screen "1000 - System" 1280x800, template "Top_Header"
   AlarmView "Alarm view_1" at 29,490 size 1237x294
   TextField "HmiScreenItemData" at 34,166 size 171x28; Text 'HMI device type:'
   TextField "HmiScreenItemData_5" at 240,166 size 299x28; Text 'TP1500 Comfort 15.0.1.0'
   TextField "HmiScreenItemData_7" at 34,199 size 171x28; Text 'Template Version:'
   TextField "HmiScreenItemData_8" at 34,263 size 171x28; Text 'Connection:'
   TextField "HmiScreenItemData_9" at 240,261 size 299x28; Text 'Simatic PLC Connection'
   TextField "HmiScreenItemData_10" at 34,293 size 171x28; Text 'PLC:'
   TextField "HmiScreenItemData_11" at 240,291 size 299x28; Text 'S7-1518F'
   TextField "HmiScreenItemData_1" at 240,199 size 299x28; Text 'FORD_Ver_1.1'
   TextField "HmiScreenItemData_12" at 34,231 size 171x28; Text 'Configuration Software:'
   TextField "HmiScreenItemData_13" at 240,229 size 299x28; Text 'WinCC TIA Portal V15 SP1'
   Button "HmiScreenItemData_4" at 29,119 size 283x41; TextOn 'System Information'; TextOff 'System Information'; PictureOn "Navigates to System information for TP1500 Comfort 14.0.1.0"; PictureOff "Navigates to System information for TP1500 Comfort 14.0.1.0"
   TextField "HmiScreenItemData_14" at 34,326 size 171x28; Text 'PLC Date / Time :'
   DateTimeField "Date/time field_2" at 238,356 size 253x36
   TextField "HmiScreenItemData_15" at 34,360 size 171x28; Text 'HMI Date / Time :'
   Button "HmiScreenItemData_2" at 622,114 size 262x48; TextOn 'System Settings'; TextOff 'System Settings'; PictureOn "Navigates to System settings for TP1500 Comfort 14.0.1.0"; PictureOff "Navigates to System settings for TP1500 Comfort 14.0.1.0"
   Button "HmiScreenItemData_6" at 29,442 size 318x44; TextOn 'System Messages'; TextOff 'System Messages'; PictureOn "Navigates to System screens for TP1500 Comfort 14.0.1.0"; PictureOff "Navigates to System screens for TP1500 Comfort 14.0.1.0"
      on Release: ActivateScreen("1000 - System", 0)
   TextField "Text field_1" at 241,328 size 48x31; Text 'Text'
   Button "Toggle language_1" at 1082,171 size 101x121; TextOn 'Toggle langu...'; TextOff 'User Admin.'
      on Release: ActivateScreen("1001 - User Adminstration", 0)
   Button "Toggle language_2" at 622,171 size 101x121; TextOn 'Toggle langu...'; TextOff 'Online'
      on Release: function_bb44b551(0)
   Button "Toggle language_3" at 736,171 size 101x121; TextOn 'Toggle langu...'; TextOff 'Offline'
      on Release: function_bb44b551(1)
   Button "Toggle language_4" at 851,171 size 101x121; TextOn 'Toggle langu...'; TextOff 'Transfer'
      on Release: function_bb44b551(2)
   Button "Toggle language_5" at 966,171 size 101x121; TextOn 'Toggle langu...'; TextOff 'Toggle Language'
      on Release: function_fb9197e8(-1)
   Button "Toggle language_6" at 622,301 size 101x121; TextOn 'Toggle langu...'; TextOff 'Calibrate Screen'
      on Release: function_bc3e350c()
   Button "Toggle language_7" at 736,301 size 101x121; TextOn 'Toggle langu...'; TextOff 'Clean Screen'
      on Release: function_be740847(30)
   Button "Toggle language_8" at 851,301 size 101x121; TextOn 'Toggle langu...'; TextOff 'Control Panel'
      on Release: function_f34a74f3()
   Button "Toggle language_9" at 965,301 size 101x121; TextOn 'Toggle langu...'; TextOff 'Stop Runtime'
      on Release: StopRuntime(0)
   Button "Toggle language_10" at 472,301 size 101x121; TextOn 'Toggle langu...'; TextOff 'Internal Software Versions'
      on Release: function_febcb963(-1)
   Button "Button_1" at 1082,301 size 102x120; TextOff 'On Screen Keyboard'
      on Release: function_d6caf649(0)
      Appearance <- "Always_OFF_HMI"

screen "1001 - User Adminstration" 1280x800, template "Top_Header"
   UserView "User view_1" at 26,185 size 1235x486
   Button "HmiScreenItemData_3" at 48,119 size 197x58; TextOn 'User Administration'; TextOff 'User Administration'; PictureOn "Navigates to User administration for TP1500 Comfort 14.0.1.0"; PictureOff "Navigates to User administration for TP1500 Comfort 14.0.1.0"

Template "TESTCENTER_SDC" 1280x800
   Button "Template_Vorlage_Schaltfläche" at 260,714 size 128x84; TextOff 'START'
      on Click: ActivateScreen("010_START", 0)
   Button "Template_Vorlage_Schaltfläche_0" at 387,714 size 128x84; TextOff 'OVERVIEW'
      on Click: ActivateScreen("700_System_Line_Overview", 0)
   Button "Template_Vorlage_Schaltfläche_1" at 514,714 size 128x84; TextOff 'TS PARAMETER'
      on Click: ActivateScreen("708_ZONE_STATUS", 0); "SDC_TS_PARAMETER"()
   Button "Template_Vorlage_Schaltfläche_2" at 641,714 size 128x84; TextOff 'EMS STATUS'
      on Click: ActivateScreen("711_CARRIER_STATUS", 0)
   Button "Template_Vorlage_Schaltfläche_3" at 768,714 size 128x84; TextOff 'Text'
   Button "Template_Vorlage_Schaltfläche_4" at 895,714 size 128x84; TextOff 'MESSAGES'
      on Click: ActivateScreen("019_MESSAGEs", 0)
   Button "Template_Vorlage_Schaltfläche_5" at 1022,714 size 128x84; TextOff 'FEHLER QUIT FAULT RESET'
      on Release: ResetBit("DB_SDC_GLOBAL_M.SDC_ER_Reset(1)")
      on Press: SetBit("DB_SDC_GLOBAL_M.SDC_ER_Reset(1)")
   Button "Template_Vorlage_Schaltfläche_6" at 1149,714 size 128x84; TextOff 'zurück / BACK'
      on Click: function_efd93a16()
   SymbolicIOField "Template_Vorlage_Symbolisches EA-Feld" at 1,3 size 671x25; TextOn '1'; TextOff '0'; TextList "SDC_ScreensName"
      ProcessValue <- "SDC\_intern_Bildnummer"
   UserView "Template_Vorlage_Vorlage_Benutzeranzeige_1" at 935,3 size 175x24
   DateTimeField "Template_Vorlage_DateTimeField_1" at 868,3 size 65x22
   DateTimeField "Template_Vorlage_DateTimeField_0" at 784,4 size 87x20
   GraphicView "Template_Vorlage_TemplateGraphicViewLogo_1" at 1112,3 size 167x25; Picture "Siemens"
   GraphicIOField "Template_Vorlage_Grafisches EA-Feld_1" at 2,4 size 20x20; PictureList "Grafikliste_G_Y"
      ProcessValue <- "Clock_1Hz"
   IOField "Vorlage_EA-Feld_2" at 754,4 size 44x19; FormatPattern 9999
      ProcessValue <- "_intern_Pult_Nr"
   TextField "Vorlage_Textfeld_1" at 677,3 size 89x23; Text 'PultNr. SDC'
   Button "Template_Vorlage_Schaltfläche_7" at 2,714 size 258x84; TextOff 'Text'
   AlarmView "Template_Vorlage_AlarmsLine_1" at 0,676 size 1280x36; ColumnTextDevice 'PLC / Steuerung / ПЛК'; ColumnTextNumber 'Nr. / No. / 编号 / № / N.º.'; ColumnTextAckGroup 'Gruppe quittieren / QGR / Acknowledge group / 确认组 / Квитировать группу / Acusar grupo'; ColumnTextAlarmState 'Status / Zustand / 状态 / Статус / Estado'; ColumnTextTime 'Zeit / Uhrzeit / Time / 时间 / Время / Hora'; ColumnTextDate 'Datum / Date / 日期 / Дата / Fecha'; ColumnTextAlarmText 'Text / 文本 / Текст / Texto'

Template "SDC" 1280x800
   SymbolicIOField "Template_Vorlage_Symbolisches EA-Feld" at 261,2 size 708x31; TextOn '1'; TextOff '0'; TextList "SDC_ScreensName"
      ProcessValue <- "SDC\_intern_Bildnummer"
   GraphicView "Template_Vorlage_TemplateGraphicViewLogo_1" at 1107,5 size 167x25; Picture "Siemens"
   GraphicIOField "Template_Vorlage_Grafisches EA-Feld_1" at 1081,8 size 20x20; PictureList "Grafikliste_G_Y"
      ProcessValue <- "Clock_1Hz"
   Button "Template_Vorlage_Schaltfläche" at 11,714 size 128x84; TextOff 'HOME / START'
      on Click: ActivateScreen("010_START", 0)
   Button "Template_Vorlage_Schaltfläche_1" at 271,714 size 128x84; TextOff 'TS PAR. TS PARAMETER'
      on Click: ActivateScreen("708_ZONE_STATUS", 0); "SDC_TS_PARAMETER"()
   Button "Template_Vorlage_Schaltfläche_2" at 401,714 size 128x84; TextOff 'EMS STATUS'
      on Click: ActivateScreen("711_CARRIER_STATUS", 0)
   Button "Template_Vorlage_Schaltfläche_4" at 888,714 size 128x84; TextOff 'ERRORS / MESSAGES / MELDUNGEN'
      on Click: ActivateScreen("019_MESSAGEs", 0)
   Button "Template_Vorlage_Schaltfläche_5" at 1018,714 size 128x84; TextOff 'QUIT FAULT RESET'
      on Release: ResetBit("DB_SDC_GLOBAL_M.SDC_ER_Reset")
      on Press: SetBit("DB_SDC_GLOBAL_M.SDC_ER_Reset")
   Button "Template_Vorlage_Schaltfläche_6" at 1148,714 size 128x84; TextOff 'BACK / ZURÜCK'
      on Click: function_efd93a16()
   Button "Template_Vorlage_Schaltfläche_3" at 141,714 size 128x84; TextOff 'GLOB. PAR. START GLOBAL PARAMETER'
      on Click: ActivateScreen("707_GLOBAL_PARAMETER", 0)
   TextField "Vorlage_Textfeld_1" at 909,6 size 127x25; Text 'DeskNo. SDC'
   IOField "Vorlage_EA-Feld_1" at 1039,4 size 41x29; FormatPattern 999
      ProcessValue <- "_intern_Pult_Nr"
   TextField "Template_Vorlage_OBJECT_3" at 1,1 size 70x32; Text 'TIME: / Zeit:'
      Appearance <- "TP_Online"
   DateTimeField "Template_Vorlage_OBJECT_5" at 56,1 size 114x32
      Appearance <- "TP_Online"
   DateTimeField "Vorlage_Datum/Uhrzeit-Feld_1" at 169,4 size 123x26

Template "Top_Header" 1280x800
   Button "Template_Button_3" at 1074,2 size 203x55; TextOn 'FAULT RESET FAULT RESET'; TextOff 'FAULT RESET FAULT RESET'
      on Release: ResetBit("DB_SDC_GLOBAL_M.SDC_ER_Reset")
      on Press: SetBit("DB_SDC_GLOBAL_M.SDC_ER_Reset")
   AlarmView "Template_Alarm view_2" at 128,2 size 948x112
   Button "Template_Button_4" at 1196,56 size 81x59; TextOff 'Text'
      Appearance <- "AlwaysTRUE"
   Button "Button_7" at 0,57 size 128x58; TextOff 'SELECT SCREEN'
      on Release: ActivateScreen("010_START", 0)
   Button "Button_6" at 0,0 size 128x58; TextOff 'PREVIOUS SCREEN'
      on Click: function_efd93a16()
   DateTimeField "Template_Date/time field_2" at 1075,56 size 123x28
   DateTimeField "Template_Date/time field_3" at 1075,83 size 122x32

PopupScreen "Pop-up_OverviewModules" 1280x800
   Button "Schaltfläche_64" at 1110,723 size 119x49; TextOn 'schließen / close'; TextOff 'schließen / close'
      on Click: function_efd93a16("Pop-up_OverviewModules", 0, 0, 0, -1, 2); ResetBit("UserDiag_HmiData_ioSlotDiagnosticsLoaded")
   IOField "I/O field_2" at 241,713 size 579x49; FormatPattern ??????????????????????????????????????????????????
      ProcessValue <- "UserDiag_HmiData_actDeviceName"
   IOField "I/O field_1" at 241,647 size 60x49; FormatPattern 999
      ProcessValue <- "actIOSystemNumber"
   IOField "I/O field_3" at 383,647 size 60x49; FormatPattern 999
      ProcessValue <- "UserDiag_HmiData_actDeviceNumber"
   TextField "Text field_1" at 137,658 size 107x26; Text 'IO System'
   TextField "Text field_2" at 314,658 size 72x26; Text 'Device'
      Visibility <- "actIOSystemNumber"
   TextField "Text field_3" at 181,724 size 62x26; Text 'Name'
   ScreenModuleView "typeSlot_1" at 67,22 size 49x152; Guid_{11997190-58737} '01'; ScreenModuleType ""
      Guid_{11997190-58740} <- "[1]"
      Guid_{11997190-58743} <- "[1]"
   ScreenModuleView "typeSlot_2" at 20,22 size 49x152; ScreenModuleType ""
      Guid_{11997190-58740} <- "[0]"
      Guid_{11997190-58743} <- "[0]"
   ScreenModuleView "typeSlot_3" at 115,22 size 49x152; Guid_{11997190-58737} '02'; ScreenModuleType ""
      Guid_{11997190-58740} <- "[2]"
      Guid_{11997190-58743} <- "[2]"
   ScreenModuleView "typeSlot_4" at 162,22 size 49x152; Guid_{11997190-58737} '03'; ScreenModuleType ""
      Guid_{11997190-58740} <- "[3]"
      Guid_{11997190-58743} <- "[3]"
   ScreenModuleView "typeSlot_5" at 210,22 size 49x152; Guid_{11997190-58737} '04'; ScreenModuleType ""
      Guid_{11997190-58740} <- "[4]"
      Guid_{11997190-58743} <- "[4]"
   ScreenModuleView "typeSlot_6" at 257,22 size 49x152; Guid_{11997190-58737} '05'; ScreenModuleType ""
      Guid_{11997190-58740} <- "[5]"
      Guid_{11997190-58743} <- "[5]"
   ScreenModuleView "typeSlot_7" at 305,22 size 49x152; Guid_{11997190-58737} '06'; ScreenModuleType ""
      Guid_{11997190-58740} <- "[6]"
      Guid_{11997190-58743} <- "[6]"
   ScreenModuleView "typeSlot_8" at 352,22 size 49x152; Guid_{11997190-58737} '07'; ScreenModuleType ""
      Guid_{11997190-58740} <- "[7]"
      Guid_{11997190-58743} <- "[7]"
   ScreenModuleView "typeSlot_9" at 400,22 size 49x152; Guid_{11997190-58737} '08'; ScreenModuleType ""
      Guid_{11997190-58740} <- "[8]"
      Guid_{11997190-58743} <- "[8]"
   ScreenModuleView "typeSlot_10" at 447,22 size 49x152; Guid_{11997190-58737} '09'; ScreenModuleType ""
      Guid_{11997190-58740} <- "[9]"
      Guid_{11997190-58743} <- "[9]"
   ScreenModuleView "typeSlot_11" at 495,22 size 49x152; Guid_{11997190-58737} '10'; ScreenModuleType ""
      Guid_{11997190-58740} <- "[10]"
      Guid_{11997190-58743} <- "[10]"
   ScreenModuleView "typeSlot_12" at 542,22 size 49x152; Guid_{11997190-58737} '11'; ScreenModuleType ""
      Guid_{11997190-58740} <- "[11]"
      Guid_{11997190-58743} <- "[11]"
   ScreenModuleView "typeSlot_13" at 590,22 size 49x152; Guid_{11997190-58737} '12'; ScreenModuleType ""
      Guid_{11997190-58740} <- "[12]"
      Guid_{11997190-58743} <- "[12]"
   ScreenModuleView "typeSlot_14" at 637,22 size 49x152; Guid_{11997190-58737} '13'; ScreenModuleType ""
      Guid_{11997190-58740} <- "[13]"
      Guid_{11997190-58743} <- "[13]"
   ScreenModuleView "typeSlot_15" at 685,22 size 49x152; Guid_{11997190-58737} '14'; ScreenModuleType ""
      Guid_{11997190-58740} <- "[14]"
      Guid_{11997190-58743} <- "[14]"
   ScreenModuleView "typeSlot_16" at 733,22 size 49x152; Guid_{11997190-58737} '15'; ScreenModuleType ""
      Guid_{11997190-58740} <- "[15]"
      Guid_{11997190-58743} <- "[15]"
   ScreenModuleView "typeSlot_17" at 780,22 size 49x152; Guid_{11997190-58737} '16'; ScreenModuleType ""
      Guid_{11997190-58740} <- "[16]"
      Guid_{11997190-58743} <- "[16]"
   ScreenModuleView "typeSlot_18" at 828,22 size 49x152; Guid_{11997190-58737} '17'; ScreenModuleType ""
      Guid_{11997190-58740} <- "[17]"
      Guid_{11997190-58743} <- "[17]"
   ScreenModuleView "typeSlot_19" at 875,22 size 49x152; Guid_{11997190-58737} '18'; ScreenModuleType ""
      Guid_{11997190-58740} <- "[18]"
      Guid_{11997190-58743} <- "[18]"
   ScreenModuleView "typeSlot_20" at 923,22 size 49x152; Guid_{11997190-58737} '19'; ScreenModuleType ""
      Guid_{11997190-58740} <- "[19]"
      Guid_{11997190-58743} <- "[19]"
   ScreenModuleView "typeSlot_21" at 971,22 size 49x152; Guid_{11997190-58737} '20'; ScreenModuleType ""
      Guid_{11997190-58740} <- "[20]"
      Guid_{11997190-58743} <- "[20]"
   ScreenModuleView "typeSlot_22" at 20,197 size 49x152; Guid_{11997190-58737} '21'; ScreenModuleType ""
      Guid_{11997190-58740} <- "[21]"
      Guid_{11997190-58743} <- "[21]"
   ScreenModuleView "typeSlot_23" at 67,197 size 49x152; Guid_{11997190-58737} '22'; ScreenModuleType ""
      Guid_{11997190-58740} <- "[22]"
      Guid_{11997190-58743} <- "[22]"
   ScreenModuleView "typeSlot_24" at 115,197 size 49x152; Guid_{11997190-58737} '23'; ScreenModuleType ""
      Guid_{11997190-58740} <- "[23]"
      Guid_{11997190-58743} <- "[23]"
   ScreenModuleView "typeSlot_25" at 162,197 size 49x152; Guid_{11997190-58737} '24'; ScreenModuleType ""
      Guid_{11997190-58740} <- "[24]"
      Guid_{11997190-58743} <- "[24]"
   ScreenModuleView "typeSlot_26" at 210,197 size 49x152; Guid_{11997190-58737} '25'; ScreenModuleType ""
      Guid_{11997190-58740} <- "[25]"
      Guid_{11997190-58743} <- "[25]"
   ScreenModuleView "typeSlot_27" at 257,197 size 49x152; Guid_{11997190-58737} '26'; ScreenModuleType ""
      Guid_{11997190-58740} <- "[26]"
      Guid_{11997190-58743} <- "[26]"
   ScreenModuleView "typeSlot_28" at 305,197 size 49x152; Guid_{11997190-58737} '27'; ScreenModuleType ""
      Guid_{11997190-58740} <- "[27]"
      Guid_{11997190-58743} <- "[27]"
   ScreenModuleView "typeSlot_29" at 352,197 size 49x152; Guid_{11997190-58737} '28'; ScreenModuleType ""
      Guid_{11997190-58740} <- "[28]"
      Guid_{11997190-58743} <- "[28]"
   ScreenModuleView "typeSlot_30" at 400,197 size 49x152; Guid_{11997190-58737} '29'; ScreenModuleType ""
      Guid_{11997190-58740} <- "[29]"
      Guid_{11997190-58743} <- "[29]"
   ScreenModuleView "typeSlot_31" at 448,197 size 49x152; Guid_{11997190-58737} '30'; ScreenModuleType ""
      Guid_{11997190-58740} <- "[30]"
      Guid_{11997190-58743} <- "[30]"
   ScreenModuleView "typeSlot_32" at 495,197 size 49x152; Guid_{11997190-58737} '31'; ScreenModuleType ""
      Guid_{11997190-58740} <- "[31]"
      Guid_{11997190-58743} <- "[31]"
   IOField "I/O field_4" at 562,647 size 60x49; FormatPattern 999
      Visibility <- "actIOSystemNumber"
      ProcessValue <- "[0]"
   TextField "Text field_4" at 452,658 size 112x26; Text 'IP Adresse / IP address'
      Visibility <- "actIOSystemNumber"
   IOField "I/O field_5" at 628,647 size 60x49; FormatPattern 999
      Visibility <- "actIOSystemNumber"
      ProcessValue <- "[1]"
   IOField "I/O field_6" at 694,647 size 60x49; FormatPattern 999
      Visibility <- "actIOSystemNumber"
      ProcessValue <- "[2]"
   IOField "I/O field_7" at 760,647 size 60x49; FormatPattern 999
      Visibility <- "actIOSystemNumber"
      ProcessValue <- "[3]"
   TextField "Text field_5" at 325,658 size 58x26; Text 'Slave'
      Visibility <- "actIOSystemNumber"

PopupScreen "Pop-up_Legend" 1280x800
   TextField "Text field_1" at 15,5 size 100x49; Text 'Legende / Legend'
   TextField "Text field_2" at 80,80 size 103x26; Text 'Status OK / State OK'
   TextField "Text field_3" at 80,146 size 165x26; Text 'Status GESTÖRT / State FAULTY'
   TextField "Text field_4" at 80,212 size 254x26; Text 'Status AUSGEFALLEN / State LOST CONNECTION'
   TextField "Text field_5" at 80,277 size 211x26; Text 'Status DEAKTIVIERT / State DEACTIVATED'
   TextField "Text field_6" at 80,343 size 339x26; Text 'Status PROBLEM / MAINTENANCE / State PROBLEM / MAINTENANCE'
   TextField "Text field_7" at 80,409 size 268x26; Text 'Status GESTÖRT GEWESEN / State WAS FAULTY'
   TextField "Text field_8" at 80,475 size 315x26; Text 'Status AUSGEFALLEN GEWESEN / State HAD LOST CONNECTION'
   TextField "Text field_9" at 80,540 size 314x26; Text 'Status DEAKTIVIERT GEWESEN / State WAS DEACTIVATED'
   TextField "Text field_10" at 80,606 size 442x26; Text 'Status PROBLEM / MAINTENANCE GEWESEN / State WAS PROBLEM / MAINTENANCE'
   Button "Schaltfläche_64" at 1110,723 size 119x49; TextOn 'schließen / close'; TextOff 'schließen / close'
      on Click: function_efd93a16("Pop-up_Legend", 0, 0, 0, -1, 2)

screen "010_START" 1280x800, template "Top_Header"
   on GenerateScreen: function_ea909784(0, U 0, '\Storage Card USB\record.csv', 2, 1, N)
   Button "Button_1" at 775,328 size 140x105; TextOn 'GLOBAL_PARAMETER GLOBAL PARAMETER'; TextOff 'GLOBAL_PARAMETER GLOBAL PARAMETER'
      on Click: ActivateScreen("707_GLOBAL_PARAMETER", 0)
   Button "Button_7" at 535,327 size 140x105; TextOn 'SECTION STATUS SECTION STATUS'; TextOff 'SECTION STATUS ZONE STATUS'
      on Click: ActivateScreen("708_ZONE_STATUS", 0)
   Button "Button_9" at 535,454 size 140x105; TextOn 'EMS STATUS EMS STATUS'; TextOff 'EMS STATUS CARRIER STATUS'
      on Click: ActivateScreen("711_CARRIER_STATUS", 0)
   Button "Button_14" at 535,198 size 140x105; TextOn 'LINE_OVERVIEW_2 LINE OVERVIEW_2'; TextOff 'LINE_OVERVIEW_2 LINE OVERVIEW'
      on Click: ActivateScreen("700_System_Line_Overview", 0)
   Button "Button_17" at 775,585 size 140x105; TextOn 'LINE_OVERVIEW_1 / MESSAGES'; TextOff 'LINE_OVERVIEW_1 FAULT MESSAGES'
      on Click: ActivateScreen("019_MESSAGEs", 0)
   Button "Button_18" at 775,454 size 140x105; TextOn 'LINE_OVERVIEW_1 PROFINET IO DIAGNOSTICS'; TextOff 'LINE_OVERVIEW_1 PROFINET IO DIAGNOSTICS'
      on Click: ActivateScreen("752_Profinet_IO_System", 0)
   Button "Button_3" at 535,585 size 140x105; TextOn 'EMS STATUS EMS STATUS'; TextOff 'EMS STATUS ALL CARRIER STATUS'
      on Click: ActivateScreen("710_ALL_CARRIER_STATUS", 0)
   Button "Button_6" at 299,198 size 140x105; TextOn 'SECTION PARAMETER SECTION PARAMETER'; TextOff 'SECTION PARAMETER SYSTEM SCREEN'
      on Click: ActivateScreen("1000 - System", 0)
   Button "Button_10" at 299,323 size 140x105; TextOn 'SECTION STATUS SECTION STATUS'; TextOff 'SECTION STATUS SYSTEM DIAGNOSTIC'
      on Release: ActivateScreen("2003 - System Diag", 0)
   Button "Button_12" at 299,450 size 140x105; TextOn 'SECTION STATUS SECTION STATUS'; TextOff 'SECTION STATUS PLC WEB SERVER INTERFACE'
      on Release: ActivateScreen("2004 - PLC Web Server Diag", 0)
   Button "Button_13" at 299,585 size 140x105; TextOn 'SECTION STATUS SECTION STATUS'; TextOff 'SECTION STATUS USER ADMIN'
      on Click: ActivateScreen("708_ZONE_STATUS", 0)
   Button "Button_5" at 775,198 size 140x105; TextOn 'LINE_OVERVIEW_2 LINE OVERVIEW_2'; TextOff 'LINE_OVERVIEW_2 ACCESS POINT LAYOUT'
      on Click: ActivateScreen("715_ACCESS_POINT_LAYOUT", 0)

screen "019_MESSAGEs" 1280x800, template "Top_Header"
   on GenerateScreen: SetTag("SDC\_intern_Bildnummer", 190)
   Button "Vorlage_Schaltfläche_19" at 387,714 size 128x84; TextOff 'alle Meldungen All Messages'
      on Click: SetTag("SDC\_intern_MELDUNGEN", 0)
      Appearance <- "SDC\_intern_MELDUNGEN"
   Button "Vorlage_Schaltfläche_20" at 514,714 size 128x84; TextOff 'Störungen / Errors'
      on Click: SetTag("SDC\_intern_MELDUNGEN", 1)
      Appearance <- "SDC\_intern_MELDUNGEN"
   Button "Vorlage_Schaltfläche_21" at 768,714 size 128x84; TextOff 'Meldungen / Reports'
      on Click: SetTag("SDC\_intern_MELDUNGEN", 3)
      Appearance <- "SDC\_intern_MELDUNGEN"
   Button "Vorlage_Schaltfläche_26" at 641,714 size 128x84; TextOff 'Warnungen / Warnings'
      on Click: SetTag("SDC\_intern_MELDUNGEN", 2)
      Appearance <- "SDC\_intern_MELDUNGEN"
   Button "Vorlage_Schaltfläche_27" at 1150,714 size 128x84; TextOff 'Archiv / Archive'
      on Click: SetTag("SDC\_intern_MELDUNGEN", 7)
      Appearance <- "SDC\_intern_MELDUNGEN"
   Button "Vorlage_Schaltfläche_22" at 895,714 size 128x84; TextOff 'Personen- schutz Personal Protection'
      on Click: SetTag("SDC\_intern_MELDUNGEN", 4)
      Appearance <- "SDC\_intern_MELDUNGEN"
   Button "Vorlage_Schaltfläche_23" at 1023,714 size 128x84; TextOff 'Bus- meldungen Bus- Messages'
      on Click: SetTag("SDC\_intern_MELDUNGEN", 5)
      Appearance <- "SDC\_intern_MELDUNGEN"
   AlarmView "Alles" at 15,121 size 1254x580; ColumnTextDevice 'PLC / Controls / ПЛК'; ColumnTextNumber 'Nr. / No. / 编号 / № / N.º.'; ColumnTextAckGroup 'Gruppe quittieren / QGR / Acknowledge group / 确认组 / Квитировать группу / Acusar grupo'; ColumnTextAlarmState 'Status / 状态 / Статус / Estado'; ColumnTextTime 'Zeit / Time / 时间 / Время / Hora'; ColumnTextDate 'Datum / Date / 日期 / Дата / Fecha'; ColumnTextAlarmText 'Text / 文本 / Текст / Texto'

screen "712_CARRIER_IO" 1280x800, template "Top_Header"
   on GenerateScreen: "SDC_EMS_STATUS"('SDC\_EMS_Nr'); "SDC_TS_REFERENCE"("SDC\_TS_Nr"); SetTag("SDC\_intern_Bildnummer", 712); "SDC_EMS_TA_STATUS"("HMI_EMS_Nr"); SetTag("SDC\_intern_Bildnummer", 712)
   on ClearScreen: SetTag("SDC\DB_SDC_EMS\HMI[XX].BILD_Nr", 0)
   IOField "EA-Feld_4" at 510,185 size 56x32; FormatPattern 9999
      on OnFinishInput: "SDC_EMS_STATUS"("HMI_EMS_Nr"); "SDC_TS_REFERENCE"("SDC\DB_SDC_EMS\EMS[XXX].TS_STAT.VAL.SEK"); "SDC_EMS_TA_STATUS"("HMI_EMS_Nr"); "SDC_ERRORS"("HMI_EMS_Nr")
      ProcessValue <- "HMI_EMS_Nr"
   TextField "Textfeld_3" at 618,188 size 118x25; Text 'EMS-No. / EMS-Number / Carrier-Number'
   Button "Schaltfläche_1" at 567,185 size 40x32; TextOff '+'
      on Click: function_dd21b452("HMI_EMS_Nr", 1); "SDC_EMS_STATUS"("HMI_EMS_Nr"); "SDC_EMS_TA_STATUS"("HMI_EMS_Nr"); "SDC_ERRORS"("HMI_EMS_Nr")
   Button "Schaltfläche_3" at 470,185 size 39x32; TextOff '-'
      on Click: function_b9b71300("HMI_EMS_Nr", 1); "SDC_EMS_STATUS"("HMI_EMS_Nr"); "SDC_EMS_TA_STATUS"("HMI_EMS_Nr"); "SDC_ERRORS"("HMI_EMS_Nr")
   TextField "Textfeld_7" at 488,118 size 243x27; Text 'section counter / min Barcode mm / Carrier I/O'
   Button "Button_1" at 92,309 size 50x432; TextOff 'Text'
   TextField "Textfeld_4" at 54,281 size 135x25; Text 'EMS-No. / EMS-Number / 8 input safety I/O'
   Button "Button_2" at 425,310 size 50x432; TextOff 'Text'
   TextField "Textfeld_5" at 330,259 size 243x27; Text 'section counter / min Barcode mm / Slot 3'
   Button "Button_3" at 710,311 size 50x432; TextOff 'Text'
   TextField "Textfeld_1" at 615,260 size 243x27; Text 'section counter / min Barcode mm / Slot 4'
   TextField "Textfeld_8" at 653,283 size 164x25; Text 'EMS-No. / EMS-Number / 16 input standard I/O'
   Button "Button_4" at 1047,311 size 50x432; TextOff 'Text'
   TextField "Textfeld_9" at 953,261 size 243x27; Text 'section counter / min Barcode mm / Slot 5'
   TextField "Textfeld_11" at 145,317 size 100x25; Text 'EMS-No. / EMS-Number / I10.0 SPARE'
   TextField "Textfeld_6" at 383,281 size 146x25; Text 'EMS-No. / EMS-Number / 8 output safety I/O'
   TextField "Textfeld_12" at 989,283 size 166x25; Text 'EMS-No. / EMS-Number / 8 output standard I/O'
   TextField "Textfeld_10" at 145,343 size 100x25; Text 'EMS-No. / EMS-Number / I10.1 SPARE'
   TextField "Textfeld_13" at 145,369 size 100x25; Text 'EMS-No. / EMS-Number / I10.2 SPARE'
   TextField "Textfeld_14" at 145,395 size 100x25; Text 'EMS-No. / EMS-Number / I10.3 SPARE'
   TextField "Textfeld_15" at 145,420 size 100x25; Text 'EMS-No. / EMS-Number / I10.4 SPARE'
   TextField "Textfeld_16" at 145,446 size 100x25; Text 'EMS-No. / EMS-Number / I10.5 SPARE'
   TextField "Textfeld_17" at 145,472 size 100x25; Text 'EMS-No. / EMS-Number / I10.6 SPARE'
   TextField "Textfeld_18" at 145,498 size 100x25; Text 'EMS-No. / EMS-Number / I10.7 SPARE'
   TextField "Textfeld_19" at 479,317 size 100x25; Text 'EMS-No. / EMS-Number / Q6.0 SPARE'
   TextField "Textfeld_20" at 479,343 size 100x25; Text 'EMS-No. / EMS-Number / Q6.1 SPARE'
   TextField "Textfeld_21" at 479,369 size 100x25; Text 'EMS-No. / EMS-Number / Q6.2 SPARE'
   TextField "Textfeld_22" at 479,395 size 100x25; Text 'EMS-No. / EMS-Number / Q6.3 SPARE'
   TextField "Textfeld_23" at 479,420 size 100x25; Text 'EMS-No. / EMS-Number / Q6.4 SPARE'
   TextField "Textfeld_24" at 479,446 size 100x25; Text 'EMS-No. / EMS-Number / Q6.5 SPARE'
   TextField "Textfeld_25" at 479,472 size 100x25; Text 'EMS-No. / EMS-Number / Q6.6 SPARE'
   TextField "Textfeld_26" at 479,498 size 100x25; Text 'EMS-No. / EMS-Number / Q6.7 SPARE'
   TextField "Textfeld_27" at 765,317 size 259x25; Text 'EMS-No. / EMS-Number / I11.0 480 VAC POWER ON MDCB1'
   TextField "Textfeld_28" at 765,344 size 196x25; Text 'EMS-No. / EMS-Number / I11.1 ACCUM. PHOTOEYE'
   TextField "Textfeld_29" at 765,370 size 100x25; Text 'EMS-No. / EMS-Number / I11.2 SPARE'
   TextField "Textfeld_30" at 765,397 size 100x25; Text 'EMS-No. / EMS-Number / I11.3 SPARE'
   TextField "Textfeld_31" at 765,422 size 210x25; Text 'EMS-No. / EMS-Number / I11.4 DC SUPPLY ON PSCB2'
   TextField "Textfeld_32" at 765,447 size 100x25; Text 'EMS-No. / EMS-Number / I11.5 SPARE'
   TextField "Textfeld_33" at 765,475 size 213x25; Text 'EMS-No. / EMS-Number / I11.6 CRASH DETECT PROX'
   TextField "Textfeld_34" at 765,501 size 100x25; Text 'EMS-No. / EMS-Number / I11.7 SPARE'
   TextField "Textfeld_35" at 765,527 size 207x25; Text 'EMS-No. / EMS-Number / I12.0 PB1 - PROD HOLD LH'
   TextField "Textfeld_36" at 765,553 size 165x25; Text 'EMS-No. / EMS-Number / I12.1 PB2 - RESET LH'
   TextField "Textfeld_37" at 765,579 size 210x25; Text 'EMS-No. / EMS-Number / I12.2 PB3 - PROD HOLD RH'
   TextField "Textfeld_38" at 765,605 size 168x25; Text 'EMS-No. / EMS-Number / I12.3 PB4 - RESET RH'
   TextField "Textfeld_39" at 765,630 size 100x25; Text 'EMS-No. / EMS-Number / I12.4 SPARE'
   TextField "Textfeld_40" at 765,656 size 100x25; Text 'EMS-No. / EMS-Number / I12.5 SPARE'
   TextField "Textfeld_41" at 765,682 size 100x25; Text 'EMS-No. / EMS-Number / I12.6 SPARE'
   TextField "Textfeld_42" at 765,708 size 100x25; Text 'EMS-No. / EMS-Number / I12.7 SPARE'
   TextField "Textfeld_43" at 1101,319 size 145x25; Text 'EMS-No. / EMS-Number / Q4.0 SITOP RESET'
   TextField "Textfeld_44" at 1101,345 size 158x25; Text 'EMS-No. / EMS-Number / Q4.1 FAULT LIGHT 1'
   TextField "Textfeld_45" at 1101,371 size 142x25; Text 'EMS-No. / EMS-Number / Q4.2 RUN LIGHT 1'
   TextField "Textfeld_46" at 1101,397 size 158x25; Text 'EMS-No. / EMS-Number / Q4.3 FAULT LIGHT 2'
   TextField "Textfeld_47" at 1101,422 size 142x25; Text 'EMS-No. / EMS-Number / Q4.4 RUN LIGHT 2'
   TextField "Textfeld_48" at 1101,448 size 100x25; Text 'EMS-No. / EMS-Number / Q4.5 SPARE'
   TextField "Textfeld_49" at 1101,474 size 100x25; Text 'EMS-No. / EMS-Number / Q4.6 SPARE'
   TextField "Textfeld_50" at 1101,500 size 100x25; Text 'EMS-No. / EMS-Number / Q4.7 SPARE'
   Circle "Kreis_13" at 110,320 size 15x15
      Appearance <- "HMI_Status_Slot2_Inputs"
   Circle "Kreis_1" at 110,344 size 15x15
      Appearance <- "HMI_Status_Slot2_Inputs"
   Circle "Kreis_2" at 110,370 size 15x15
      Appearance <- "HMI_Status_Slot2_Inputs"
   Circle "Kreis_3" at 110,396 size 15x15
      Appearance <- "HMI_Status_Slot2_Inputs"
   Circle "Kreis_4" at 110,422 size 15x15
      Appearance <- "HMI_Status_Slot2_Inputs"
   Circle "Kreis_5" at 110,448 size 15x15
      Appearance <- "HMI_Status_Slot2_Inputs"
   Circle "Kreis_6" at 110,474 size 15x15
      Appearance <- "HMI_Status_Slot2_Inputs"
   Circle "Kreis_7" at 110,500 size 15x15
      Appearance <- "HMI_Status_Slot2_Inputs"
   Circle "Kreis_17" at 443,319 size 15x15
      Appearance <- "HMI_Status_Slot3_Outputs"
   Circle "Kreis_18" at 443,345 size 15x15
      Appearance <- "HMI_Status_Slot3_Outputs"
   Circle "Kreis_19" at 443,371 size 15x15
      Appearance <- "HMI_Status_Slot3_Outputs"
   Circle "Kreis_20" at 443,397 size 15x15
      Appearance <- "HMI_Status_Slot3_Outputs"
   Circle "Kreis_21" at 443,423 size 15x15
      Appearance <- "HMI_Status_Slot3_Outputs"
   Circle "Kreis_22" at 443,449 size 15x15
      Appearance <- "HMI_Status_Slot3_Outputs"
   Circle "Kreis_23" at 443,475 size 15x15
      Appearance <- "HMI_Status_Slot3_Outputs"
   Circle "Kreis_24" at 443,501 size 15x15
      Appearance <- "HMI_Status_Slot3_Outputs"
   Circle "Kreis_33" at 728,320 size 15x15
      Appearance <- "HMI_Status_Slot4_Inputs"
   Circle "Kreis_34" at 728,346 size 15x15
      Appearance <- "HMI_Status_Slot4_Inputs"
   Circle "Kreis_35" at 728,372 size 15x15
      Appearance <- "HMI_Status_Slot4_Inputs"
   Circle "Kreis_36" at 728,398 size 15x15
      Appearance <- "HMI_Status_Slot4_Inputs"
   Circle "Kreis_37" at 728,424 size 15x15
      Appearance <- "HMI_Status_Slot4_Inputs"
   Circle "Kreis_38" at 728,450 size 15x15
      Appearance <- "HMI_Status_Slot4_Inputs"
   Circle "Kreis_39" at 728,476 size 15x15
      Appearance <- "HMI_Status_Slot4_Inputs"
   Circle "Kreis_40" at 728,502 size 15x15
      Appearance <- "HMI_Status_Slot4_Inputs"
   Circle "Kreis_41" at 728,528 size 15x15
      Appearance <- "HMI_Status_Slot4_Inputs"
   Circle "Kreis_42" at 728,554 size 15x15
      Appearance <- "HMI_Status_Slot4_Inputs"
   Circle "Kreis_43" at 728,580 size 15x15
      Appearance <- "HMI_Status_Slot4_Inputs"
   Circle "Kreis_44" at 728,606 size 15x15
      Appearance <- "HMI_Status_Slot4_Inputs"
   Circle "Kreis_45" at 728,632 size 15x15
      Appearance <- "HMI_Status_Slot4_Inputs"
   Circle "Kreis_46" at 728,658 size 15x15
      Appearance <- "HMI_Status_Slot4_Inputs"
   Circle "Kreis_47" at 728,684 size 15x15
      Appearance <- "HMI_Status_Slot4_Inputs"
   Circle "Kreis_48" at 728,708 size 15x15
      Appearance <- "HMI_Status_Slot4_Inputs"
   Circle "Kreis_49" at 1065,320 size 15x15
      Appearance <- "HMI_Status_Slot5_Outputs"
   Circle "Kreis_50" at 1065,346 size 15x15
      Appearance <- "HMI_Status_Slot5_Outputs"
   Circle "Kreis_51" at 1065,372 size 15x15
      Appearance <- "HMI_Status_Slot5_Outputs"
   Circle "Kreis_52" at 1065,398 size 15x15
      Appearance <- "HMI_Status_Slot5_Outputs"
   Circle "Kreis_53" at 1065,424 size 15x15
      Appearance <- "HMI_Status_Slot5_Outputs"
   Circle "Kreis_54" at 1065,450 size 15x15
      Appearance <- "HMI_Status_Slot5_Outputs"
   Circle "Kreis_55" at 1065,476 size 15x15
      Appearance <- "HMI_Status_Slot5_Outputs"
   Circle "Kreis_56" at 1065,502 size 15x15
      Appearance <- "HMI_Status_Slot5_Outputs"
   TextField "Textfeld_2" at 54,259 size 125x27; Text 'section counter / min Barcode mm / Slot 2'